// TIA Portal project "g" (V14) (continued)

   REGION Init
       IF #mb_query.z.run.state = #INIT_QUERY THEN
           // Modicon convention address conversion.
           "mb_internal_a"(mode104 := false,
                          Mode => #master.MODE,
                          Data_addr => #master.DATA_ADDR,
                          mb_query := #mb_query);
           // Copy buffer to a non optimiced memory area.
           IF #mb_query.z.run.write THEN
               #buffer.buffer := #mb_query.z.buffer;
           END_IF;
           // Automatically adjust timeout.
           #comm_load.RESP_TO := T_CONV
           (* *)("mb_timeout_rtu_calc"
                 (**)(gain := #conf.timeout_gain, 
                 (**) offset := #conf.timeout_offset,
                 (**) baud := #baud, mb_query := #mb_query));
           #comm_load.RETRIES := #conf.retries;
       END_IF;

       // Initiate the hardware
       #comm_load(REQ := #mb_query.z.run.state = #INIT_QUERY,
                  PORT := #hardware_id,
                  BAUD := #baud,
                  PARITY := #conf.parity, // Even is default.
                  RESP_TO := #comm_load.RESP_TO,
                  MB_DB := #master);

       IF #mb_query.z.run.state = #INIT_QUERY THEN
           IF #comm_load.DONE THEN
               #mb_query.z.run.state := #EXEC_QUERY;
           ELSE
               // Skip query exec. if init hw didn't go well.
               // The state RECIVE_RESUALT is inside mb_query.
               #mb_query.z.run.state := #RECIVE_RESUALT;
               #mb_query.stat.done := false;
               #mb_query.stat.error := true;
               #mb_query.stat.error_comm := true;
               #mb_query.stat.status := #comm_load.STATUS;
           END_IF;
       END_IF;
   END_REGION

   REGION Exec
       // The core master block.
       #master(REQ := #mb_query.z.run.state = #EXEC_QUERY
               AND NOT #master.BUSY,
               MB_ADDR := #mb_query.z.q.mb_addr,
               MODE := #master.MODE,
               DATA_ADDR := #master.DATA_ADDR,
               DATA_LEN := #mb_query.z.q.data_len,
               BUSY => #mb_query.stat.busy,
               DATA_PTR := #buffer.buffer);

       IF #mb_query.z.run.state = #EXEC_QUERY THEN
           #mb_query.stat.error := #master.ERROR;
           #mb_query.stat.done := #master.DONE;
           #mb_query.stat.status := #master.STATUS;
           "mb_internal_f"(buffer := #buffer, mb_query := #mb_query);
       END_IF;
   END_REGION

   // End is a comman FB for both tcp and rtu.
   #end(mb_query := #mb_query, Error => #Error);
END_FUNCTION_BLOCK

// folder: Library/Modbus/Core/Special

FUNCTION_BLOCK "mb_delay"   // FB11, SCL
{ S7_Optimized_Access := 'TRUE' }
VERSION : 0.1
   VAR_INPUT
      delay : Time;
   END_VAR
   VAR_IN_OUT
      mb_query : "mb_query";
   END_VAR
   VAR
      "timer" : TON_TIME;
      halt : Bool;
   END_VAR
BEGIN
   // For use with modbus tcp, so the client dosen't jam a network.
   // The function halt execution of queries for a certain time

   #mb_query.z.run.qid_cnt += 1;  // The timer occupy one qid.

   IF #halt // If the timer has been activated.
       OR #delay = T#0s // #delay = T#0s => Disable function
   THEN
       PRESET_TIMER(PT := #delay, TIMER := #"timer");
       #"timer"(IN := #delay <> T#0s, PT := #delay);
       IF #"timer".Q OR #delay = T#0s THEN
           IF #halt THEN
               #mb_query.conf.halt := #halt := false; // Continue exec.
               RESET_TIMER(#"timer");
           END_IF;
           #mb_query.z.run.qid += BOOL_TO_UINT
           (* *)(#mb_query.z.run.qid = #mb_query.z.run.qid_cnt);
       END_IF;

   ELSIF #mb_query.z.run.qid_cnt = #mb_query.z.run.qid THEN
       #mb_query.conf.halt := #halt := true; // Halt exec.
   END_IF;
END_FUNCTION_BLOCK

FUNCTION_BLOCK "mb_delay_between_queries"   // FB13, SCL
{ S7_Optimized_Access := 'TRUE' }
VERSION : 0.1
   VAR_INPUT
      delay : Time;
   END_VAR
   VAR_IN_OUT
      mb_query : "mb_query";
   END_VAR
   VAR
      "timer" : TON_TIME;
      halt : Bool;
      old_state : UInt;
   END_VAR
   VAR CONSTANT
      ORIGIN : USInt := 0;
   END_VAR
BEGIN
   // For use with modbus tcp, so the client dosen't jam a network.
   // The function halt execution of queries for a certain time
   // not just once, but between every query. There should only be
   // one of this block for each client.

   IF #halt // Is exec. halted?
       OR #delay = T#0s // #delay = T#0s => Disable function.
   THEN
       PRESET_TIMER(PT := #delay, TIMER := #"timer");
       #"timer"(IN := #delay <> T#0s, PT := #delay);
       IF #"timer".Q
           OR #delay = T#0s AND #halt
       THEN
           RESET_TIMER(#"timer");
           #mb_query.conf.halt := #halt := false; // Continue exec.
       END_IF;

   ELSIF #mb_query.z.run.state <> #old_state
       AND #mb_query.z.run.state <> #ORIGIN
   THEN
       // Halt exec. when next query is about to be inserted,
       // but current query will still finish.
       #mb_query.conf.halt := #halt := true; // Halt exec.
   END_IF;
   #old_state := #mb_query.z.run.state;
END_FUNCTION_BLOCK

FUNCTION "mb_query_bits" : Void   // FC9, SCL
{ S7_Optimized_Access := 'TRUE' }
VERSION : 0.1
   VAR_IN_OUT
      data_ptr : Array[*] of Bool;
      mb_query : "mb_query";
   END_VAR
   VAR_TEMP
      discrete : Bool;
      dommy : Bool;
      lower : DInt;
      upper : DInt;
      bits : UInt;
      bytes : UDInt;   // bytes
   END_VAR
   VAR CONSTANT
      INIT_QUERY : USInt := 2;
      RECIVE_RESUALT : USInt := 4;
   END_VAR
BEGIN
   // This function may be used when the number of bits dosen't
   // add up to whole bytes, for function codes: 1, 2, 5 and 15. 
   // 
   // data_ptr need to be a one dimensional array of bools.
   // --- --- ---

   REGION Header
       IF #mb_query.z.run.qid_cnt + 1 <> #mb_query.z.run.qid
           OR #mb_query.stat.busy
       THEN
           // Skip query, qid will not match qid_cnt and
           // my_query will return.
           #mb_query(data_ptr := #dommy);
           RETURN;
       END_IF;
   END_REGION

   REGION Pre-calc
       // Some preparing calculations.
       CASE #mb_query.mode OF // A discrete query ?
           1, 2, 5, 15:
               #discrete := true;
           200..202:
               CASE #mb_query.data_addr OF
                   1..19999: // 1..9999, 10001..19999
                       #discrete := true;
               END_CASE;
       END_CASE;
       #lower := LOWER_BOUND(ARR := #data_ptr, DIM := 1);
       #upper := UPPER_BOUND(ARR := #data_ptr, DIM := 1);
       #bits := DINT_TO_UINT(#upper - #lower + 1); // Elements in array.

       // Auto data len ?
       IF #mb_query.data_len = #mb_query.c.auto_len THEN
           #bytes := (#bits + 7) / 8; // CEIL()
           #mb_query.data_len := SEL(G := #discrete,
                                     IN0 := (#bits + 15) / 16, // CEIL()
                                     IN1 := #bits);
       ELSE
           #bytes := SEL(G := #discrete,
                         IN0 := #mb_query.data_len * 2, // 1 word -> 2 bytes
                         IN1 := (#mb_query.data_len + 7) / 8); // CEIL()
       END_IF;
   END_REGION

   REGION Run
       // Disable buf.h. inside mb_query.
       #mb_query.conf.buffer_handler := false;

       // Run the query.
       #mb_query(data_ptr := #dommy);

       #mb_query.conf.buffer_handler := true; // Enable buf.h. again.
       #mb_query.data_len := #mb_query.c.auto_len; // Back to auto.
   END_REGION

   REGION Insert & recive
       IF #mb_query.z.run.state = #INIT_QUERY  // Insert query.
           AND #mb_query.z.run.write
       THEN
           // Copy the content from data_ptr to the buffer.
           GATHER_BLK(IN := #data_ptr[#lower],
                      COUNT_OUT := #bytes,
                      OUT => #mb_query.z.buffer[0]);

       ELSIF  #mb_query.Done // The query above.
           AND NOT #mb_query.z.run.write  // A read query
       THEN
           // Copy the content from the buffer to data_ptr.
           SCATTER_BLK(IN := #mb_query.z.buffer[0],
                       COUNT_IN := #bytes,
                       OUT => #data_ptr[#lower]);
       END_IF;
   END_REGION
END_FUNCTION

// folder: Library/Modbus/Core/sb

FUNCTION "mb_station_block_header" : Void   // FC10, SCL
{ S7_Optimized_Access := 'TRUE' }
VERSION : 1.0
   VAR_IN_OUT
      sb : "mb_station_block_udt";
      mb_query : "mb_query";
   END_VAR
   VAR CONSTANT
      ORIGIN : USInt := 0;
   END_VAR
BEGIN
   // Rexhip - Extended modbus library.
   // Read the top section of mb_query for more documentation.

   // Skip everything !
   IF #sb.conf.skip_code THEN
       RETURN;
   END_IF;

   #mb_query.data_len := 0; // Default is auto-length.
   #mb_query.conf.buffer_handler := true;

   // If device blocks are executeded in diffrent order, a wide wind
   // up effect will occur, (in same OB) this will prevent that.
   IF #mb_query.z.sb.reset THEN
       #sb.z.header_qid := #mb_query.z.run.qid_cnt + 1;
   END_IF;

   // Device id cnt. The first device has id "1". Increased in every
   // mb_device_header, reseted in mb_client_ctrl or mb_master_ctrl.
   #mb_query.z.sb.sid_cnt += 1;

   // mb_query set the same bellow variables to true, at insert or recive.
   // This informastion is later used at the footer.
   #mb_query.z.sb.head_insert := false;
   #mb_query.z.sb.head_recive := false;

   // Reset order, a variable that makes queries in a sb execute in order.
   // #mb_query.z.sb.order := false;

   // When #mb.mb.q.qid = #mb.mb.run.qid_cnt => "This" device has the
   // query-token !
   // - If the query-token points at this device header, or it point to a
   //   query in the previous device, that is surrounded by a if-statement
   //   and the statement is now false.
   // - A gid change can only be done if not "busy", this is to avoid a
   //   resualt from one query being intercepted by another
   IF #mb_query.z.run.qid > #mb_query.z.run.qid_cnt
       AND #mb_query.z.run.qid <= #sb.z.header_qid
       AND NOT #mb_query.stat.busy
   THEN
       // Reset.
       // Go back to the first state in mb_query. New query param. will
       // owerwrite old once.
       #mb_query.z.run.state := #ORIGIN;

       // At first the offset_qid points at the first query of this
       // device. When it has executed the offset will point at the
       // second query. When all queries has executed the offset will
       // be reset back to the first query. (footer) 
       #mb_query.z.run.qid :=
       (* *)#sb.z.header_qid + #sb.z.offset_qid;

       // Order is a variable that makes queries in sb execute in order.
       //    #mb_query.z.sb.order := true;
   END_IF;

   // - The code below is reduce the impact of setting a if-statement
   //   around queries, by setting the qid_cnt to a fixed value at this 
   //   point.
   // - mb_station_block_header will occupy one query-id.  
   #sb.z.header_qid :=
   MAX(IN1 := #mb_query.z.run.qid_cnt + 1,
       IN2 := #sb.z.header_qid);
   #mb_query.z.run.qid_cnt := #sb.z.header_qid;
END_FUNCTION

FUNCTION "mb_station_block_footer" : Void   // FC11, SCL
{ S7_Optimized_Access := 'TRUE' }
VERSION : 1.0
   VAR_IN_OUT
      sb : "mb_station_block_udt";
      mb_query : "mb_query";
   END_VAR
   VAR_TEMP
      "e" : Int;
      err : Bool;
   END_VAR
   VAR CONSTANT
      INSERT_QUERY : USInt := 1;
   END_VAR
BEGIN
   // Rexhip - Extended modbus library.
   // Read the top section of mb_query for more documentation.

   // Skip everything !
   IF #sb.conf.skip_code THEN
       RETURN;
   END_IF;

   REGION Recive
       IF #mb_query.z.sb.head_recive THEN
           // If there is a query that bellong to this device that has
           // recvied a resault. (with or without error)

           // Counter for exec. queries inside this station block.
           // Default is 1 query for each loop, but may be changed.
           #sb.z.exec_cnt += 1;

           // If this is the first succesfylly query after communication error,
           // then log the time this happen. (also exceptions)
           IF #sb.out.error_comm AND (
               #mb_query.stat.done
               OR #mb_query.stat.error AND NOT #mb_query.stat.error_comm)
           THEN
               #"e" := RD_LOC_T(#sb.log.connected_time);
           END_IF;

           IF #mb_query.stat.error THEN // Logging - failed query        
               // Store the values for debugging. data_addr will indicate witch 
               // query caused the error, and the status is indicate the error type.
               #sb.log.error_status := #mb_query.stat.status;
               #sb.log.error_data_addr := #mb_query.z.sb.log_data_addr;

               // Two counters, one for comm.error and for all other errors.
               IF #mb_query.stat.error_comm THEN
                   #sb.log.error_comm_cnt += 1; // Eg. Bad CRC, parity, etc.
               ELSE
                   #sb.log.error_exception_cnt += 1;
               END_IF;

               // Increase communication error counter. if it's a comm.error.
               // then reset the counter.  
               IF #mb_query.stat.error_comm THEN
                   #sb.z.comm_err_cnt += BOOL_TO_USINT(#sb.z.comm_err_cnt < 255);
               ELSE
                   #sb.z.comm_err_cnt := 0;
               END_IF;

               // The error_comm flag is set if x repeating comm.errors occurres.
               #err := #sb.z.comm_err_cnt > #sb.conf.max_comm_error;
               IF #err AND NOT #sb.out.error_comm THEN
                   // Log the time when the flag is set.
                   #"e" := RD_LOC_T(#sb.log.disconnected_time);
               END_IF;
               #sb.out.error_comm := #err;

               // A comm.error will not be displayed before the
               // communication_error flag is set. Other errors will be
               // diplayed once. (NOT comm.error -> normal error)
               #sb.out.error := #sb.out.error OR NOT #mb_query.stat.error_comm
               OR #sb.out.error_comm;

               // err_hold makes the error flag stay true for more then just
               // one plc-scan.
               #sb.z.err_hold := #sb.out.error;

           ELSIF #mb_query.stat.done THEN // Logging successfully query        
               #sb.log.done_cnt += 1;
               // One successfully query -> reset fault.
               #sb.out.error_comm := false;
               #sb.z.comm_err_cnt := 0;
           END_IF;

           // - If it's this devices has the retry token, (sid_retry = sid_cnt)
           //   a retry has been executed and faild. Then set the retry_finished
           //   flag.
           // - The retry-token will be passed on to the next device with
           //   communication problems when the query loop has reach
           //   the end. (Inside the mb_internal_e)
           // - The library make sure that only one station block with comm.
           //   problems will do retry for each query loop revolution. 
           #mb_query.z.sb.retry_finished :=
           #mb_query.z.sb.sid_retry = #mb_query.z.sb.sid_cnt
           AND #mb_query.stat.error_comm;

           // Only one query in the SB is executed (default). The purpose is
           // to avoid a SB with many queries to occupy the bus for long periodes
           // of time. offset_qid is incread by one when a query has executed
           // given last query didn't resualt in a timeout.
           #sb.z.offset_qid += BOOL_TO_UINT(NOT #mb_query.stat.error_comm);
       END_IF;
   END_REGION

   REGION Middle
       // If all queries for this device has been executed,
       // then reset offset_qid back to the first query.
       IF #sb.z.offset_qid >
           #mb_query.z.run.qid_cnt - #sb.z.header_qid
       THEN
           #sb.z.offset_qid := 1;

           // Also reset error falg, if the last query was successfully.
           IF NOT #sb.z.err_hold THEN
               #sb.out.error := false;
           END_IF;
           #sb.z.err_hold := false;
       END_IF;

       // If the retry-token point at this device (sid_retry=sid_cnt), and there is
       // no communication problems then pass on the retry-token to the next device.
       // The retry token tell which device with communication problem that should
       // retry establish communication.
       #mb_query.z.sb.sid_retry +=
       BOOL_TO_UINT(#mb_query.z.sb.sid_retry = #mb_query.z.sb.sid_cnt
                    AND NOT #sb.out.error_comm);
   END_REGION

   REGION Finnish
       // Several condition that resault in passing on the query-token on to the
       // next device. Skipping all or the rest of the queries for this device:              
       #sb.out.finnish :=
       #mb_query.z.sb.head_recive AND ( // Skip rest of the queries if: ->
       (* *)#sb.z.exec_cnt >= #sb.conf.exec_x_quries // Some queries has executed,
       (*           *)// wait for the next loop for the remaining queries.
       (*      *)OR #mb_query.stat.error_comm) // A query resualting in comm.error    
       OR #mb_query.z.sb.head_insert AND ( // Erase a already inserted query if: ->
       (* *)#sb.out.error_comm // This station has allready comm. problems.
       (*      *)// And, it isn't this devies turn to try again.
       (*      *)AND (#mb_query.z.sb.sid_retry <> #mb_query.z.sb.sid_cnt
       (*           *)// Or, there has allready been a retry attempt on this loop.
       (*           *)OR #mb_query.z.sb.retry_finished) // (reseted in mb_internal_e)     
       (* *)OR #sb.conf.disable    
       (* *)OR #sb.conf.exec_x_quries = 0 // Zero => disable station block.
       (* *)OR #sb.conf.read_only // The read_only flag is set, and it's a write query.
       (*      *)AND #mb_query.z.run.write);

       IF #sb.out.finnish THEN // Reset
           // Go back to the first state in mb_query. New query param. will owerwrite 
           // old once.
           #mb_query.z.run.state := #INSERT_QUERY;
           // Set to qid to the next station block.
           #mb_query.z.run.qid := #mb_query.z.run.qid_cnt + 1;
           #sb.z.exec_cnt := 0;
       END_IF;
   END_REGION
END_FUNCTION

// folder: Library/Modbus/Core/z Internal

FUNCTION_BLOCK "mb_internal_b"   // FB6, SCL
{ S7_Optimized_Access := 'FALSE' }
VERSION : 0.1
   VAR
      buffer : Array[0..249] of Byte;
   END_VAR
BEGIN
   (*
   - Buffer for mb_master and modbus_master. (modbus rtu)
   - This block has optimize data access disabled.
   - For RTU, please do not delete the even there is no code bellow.
   - This block isn't needed for modbus tcp.
   *)
END_FUNCTION_BLOCK

FUNCTION_BLOCK "mb_internal_e"   // FB7, SCL
{ S7_Optimized_Access := 'TRUE' }
VERSION : 0.1
   VAR_OUTPUT
      Error : Bool;
   END_VAR
   VAR_IN_OUT
      mb_query : "mb_query";
   END_VAR
   VAR
      err_hold : Bool;
   END_VAR
   VAR CONSTANT
      INSERT_QUERY : USInt := 1;
      EXEC_QUERY : USInt := 3;
      RECIVE_RESUALT : USInt := 4;
   END_VAR
BEGIN
   // Internal function - common for both rtu and tcp.

   // Move on to next state when query is finnished.
   IF #mb_query.z.run.state = #EXEC_QUERY 
       AND (#mb_query.stat.error OR #mb_query.stat.done)
   THEN
       #mb_query.z.run.state := #RECIVE_RESUALT;
   END_IF;


   // Anti wind up effect for qid. msg. to devices that they should
   // reset if qid grow bigger then 60000. (See mb_station_block_header)
   #mb_query.z.sb.reset := false;
   IF #mb_query.z.run.qid > 60000 THEN
       #mb_query.z.sb.reset := true;
   END_IF;

   // #error will be keeped true as long there is at least one query that
   // generate a error. 
   IF #mb_query.stat.error THEN
       #Error := true;
       #err_hold := true;
   END_IF;

   // If all queries has been executed,
   IF #mb_query.z.run.qid > #mb_query.z.run.qid_cnt THEN

       // Error handeling (see above)
       IF NOT #err_hold THEN
           #Error := false;
       END_IF;
       #err_hold := false;

       // Start over again on the first query.
       #mb_query.z.run.qid := 1;

       // The retry-id is the device that get to have retry to restoring
       // communication after the error_comm flag is set for the station.
       // When one query loop has occurred the retry id is incremented. 
       #mb_query.z.sb.sid_retry := #mb_query.z.sb.sid_retry + 1;

       // retry_finished is set after one retry has taken place. 
       // The station that has the retry-token only has one try to make 
       // successfully query.
       #mb_query.z.sb.retry_finished := false;
       IF #mb_query.z.sb.sid_retry > #mb_query.z.sb.sid_cnt THEN
           #mb_query.z.sb.sid_retry := 1;
       END_IF;

       // Station id: (not in use)
       #mb_query.z.sb.sid := #mb_query.z.sb.sid + 1;
       IF #mb_query.z.sb.sid > #mb_query.z.sb.sid_cnt THEN
           #mb_query.z.sb.sid := 1;
       END_IF;
   END_IF;

   #mb_query.z.run.qid_cnt := 0; // (Incremented in mb_query)
   #mb_query.z.sb.sid_cnt := 0; // (Incremented in mb_station_block_header)
END_FUNCTION_BLOCK

FUNCTION "mb_internal_f" : Void   // FC2, SCL
{ S7_Optimized_Access := 'TRUE' }
VERSION : 0.1
   VAR_IN_OUT
      buffer : "mb_internal_b";
      mb_query : "mb_query";
   END_VAR
   VAR_TEMP
      comm_error : Bool;
   END_VAR
BEGIN
   // Internal function - master footer

   IF #mb_query.stat.error THEN
       // Figur out if it's a communication error.
       // (Handled different from other errors)
       CASE WORD_TO_UINT(#mb_query.stat.status) OF
           16#80C8, // Timeout
           16#80E1, // Parity error
           16#80E2, // Framing error
           16#8380: // Bad CRC 
               #comm_error := true;
       END_CASE;

   ELSIF #mb_query.stat.done // Successful query
       AND NOT #mb_query.z.run.write // A read query.
   THEN
       #mb_query.z.buffer := #buffer.buffer;
   END_IF;

   #mb_query.stat.error_comm :=
   (* *)#mb_query.stat.error AND #comm_error;
END_FUNCTION

FUNCTION "mb_internal_a" : Void   // FC4, SCL
{ S7_Optimized_Access := 'TRUE' }
VERSION : 0.1
   VAR_INPUT
      mode104 : Bool;
   END_VAR
   VAR_OUTPUT
      Mode : USInt;
      Data_addr : UDInt;
   END_VAR
   VAR_IN_OUT
      mb_query : "mb_query";
   END_VAR
BEGIN
   // Internal function

   // Modicon convention address.
   #Mode := 0;
   CASE #mb_query.z.q.mode OF
       1:  // Read output bits
           #Data_addr := 1 + #mb_query.z.q.data_addr;
       2:  // Read input bits
           #Data_addr := 10001 + #mb_query.z.q.data_addr;
       3:  // Read holding reg.
           #Data_addr := 400001 + #mb_query.z.q.data_addr;
       4:  // Read input word
           IF #mode104 THEN
               #Mode := 104;
               #Data_addr := #mb_query.z.q.data_addr;
           ELSE
               #Data_addr := 30001 + #mb_query.z.q.data_addr;
           END_IF;
       5:  // Writing a single output bit
           #Mode := 1;
           #Data_addr := 1 + #mb_query.z.q.data_addr;
       6:  // Writing a single holding register
           #Mode := 1;
           #Data_addr := 400001 + #mb_query.z.q.data_addr;
       15: // Writing multiple output bits
           #Mode := 2;
           #Data_addr := 1 + #mb_query.z.q.data_addr;
       16: // Writing multiple holding registers
           #Mode := 2;
           #Data_addr := 400001 + #mb_query.z.q.data_addr;
       200..202: // Read and write
           #Mode := #mb_query.z.q.mode - 200;
           #Data_addr := #mb_query.z.q.data_addr;
       ELSE
           #Mode := #mb_query.z.q.mode;
           #Data_addr := #mb_query.z.q.data_addr;
   END_CASE;
END_FUNCTION

FUNCTION "mb_timeout_rtu_calc" : Time   // FC5, SCL
{ S7_Optimized_Access := 'TRUE' }
VERSION : 0.1
   VAR_INPUT
      gain : Real;
      offset : Time;
      baud : UDInt;
   END_VAR
   VAR_IN_OUT
      mb_query : "mb_query";
   END_VAR
   VAR_TEMP
      t : Time;
   END_VAR
BEGIN
   // Automatically adjust timeout for modbus rtu.

   IF #gain = 0 THEN
       #t := #offset;
   ELSE
       #t := T_CONV
       (REAL_TO_UINT
        (
         11000 * ( //  11: Bits: start, data, parity, stop. 
         (* *)//   * 1000: Seconds to milliseconds
         (* *)19 // Bytes: Req: mb_addr, fc, data_addr(2), data_len(2), crc(2), 
         (* *) //        + res: mb_addr, fc, byte-count, crc(2), 
         (* *) //        + start-stop -> 6 (ca 2 x 28 bits)
         (* *)+ UINT_TO_REAL(#mb_query.z.q.data_len) *
         (*     *)SEL(G := #mb_query.z.run.discrete,
                      (* *)IN0 := INT_TO_REAL(2), // Each word is to bytes.
                      (* *)IN1 := 0.125) // Eight bits in one byte. (1/8 = 0.125)
         )
         / UDINT_TO_REAL(#baud) // High baud-rate -> low timeout
         * #gain // Safty margin
         + UDINT_TO_UINT(T_CONV(#offset))
        ));
   END_IF;

   #mb_timeout_rtu_calc :=
   LIMIT(MN := T#5ms, // A least 5ms, else comm_load will throw a error.
         IN := #t,
         MX := T#65s);
END_FUNCTION

// ===== library types =====

TYPE "timerUdt"
   STRUCT
      pt : Real;   // Preset time
      format : SInt := 2;   // 1=ms, 2=sec, 3=min, 4=h, 5=day
      RT : Real;   // Remaining time
   END_STRUCT;
END_TYPE

TYPE "ioGlobalUdt"
   STRUCT
      ackAllAlarms : Bool;   // Acknowledge all alarms
      disableAllSim : Bool;   // Disable all simulation of input values
      hmiShowTags : Bool;
      _ : Bool;
      totalActiveSim : UInt;   // Total active simulations
      totalActiveAlarms : UInt;   // Total active alarms
      totalUnacknowledgedAlarms : UInt;
      totalErrors : UInt;
   END_STRUCT;
END_TYPE

TYPE "alarmRealUdt"
   STRUCT
      value : Real;
      action : SInt;
      lim : Real;   // Alarm limit
      hyst : Real;   // Hysteresis
      delay : Time;   // Alarm delay
      delayEt : Time;   // delay elapsed time
      enable : Bool;   // Enable alarm
      autoAck : Bool := TRUE;   // manual acknowledge
      dobleAck : Bool;
      ack : Bool;   // acknowledge alarm
      memAck : Bool;   // Can be used for buzzer
      Q : Bool;   // output
   END_STRUCT;
END_TYPE

TYPE "analogInUdt"
   STRUCT
      filterConst : Real;   // 0=off , const for average filter.
      unitInterval : Real;   // 00.0 to 1.00 , (raw value, after running avg filter)
      sim : Bool;   // Simulate value
      forceInsideScale : Bool := true;   // Eg. in case of more then 20mA or less then 4mA.
      Error : Bool;   // Input signal out of range.
      zOldError : Bool;   // Internal variable
      ErrorTime : DTL;   // Time when the error occurred.
      errorAction : SInt := 100;   // [%]
      scaleMin : Real := 0.0;   // Scaled value for 4mA.
      scaleMax : Real := 100.0;   // Scaled value for 20mA.
      gain : Real := 1.0;   // Muliplied with the scaled value.
      offset : Real := 0.0;   // Added to "Q".
      Q : Real;   // value
   END_STRUCT;
END_TYPE

TYPE "analogInAndAlarmsUdt"
   STRUCT
      ai : "analogInUdt";
      execAiLogic : Bool := true;
      alarmL : "alarmRealUdt";
      alarmLL : "alarmRealUdt";
      alarmH : "alarmRealUdt";
      alarmHH : "alarmRealUdt";
      hmi : Struct
         copyAllSettings : Bool;
         pasteAllSettings : Bool;
         showTag : Bool;
      END_STRUCT;
   END_STRUCT;
END_TYPE

TYPE "alarmBoolSimpleUdt"
   STRUCT
      in : Bool;   // Input
      enable : Bool;   // Enable alarm
      autoAck : Bool := TRUE;   // Alarm will go away automaticaly when in goes false.
      dobleAck : Bool;
      ack : Bool;   // Acknowledge alarm
      memAck : Bool;   // Active alarm has been acknowledged
      Q : Bool;   // Output
   END_STRUCT;
END_TYPE

TYPE "digitalInUdt"
   STRUCT
      sim : Bool;   // Simulate input
      invert : Bool;   // Invert input
      Error : Bool;   // External error
      Q : Bool;   // Output
      delay : Time;   // Input delay
      delayEt : Time;
      alarm : "alarmBoolSimpleUdt";
      timeOn : DTL;
      timeOff : DTL;
   END_STRUCT;
END_TYPE

TYPE "intervalUdt"
   STRUCT
      time_between : Real;
      time_active : Real;
      time_format : SInt := 2;   // 1=ms, 2=sec, 3=min, 4=h, 5=day
      force_on : Bool;
      force_off : Bool;
      Q : Bool;
      RT : Real;
   END_STRUCT;
END_TYPE

TYPE "load_balancer_info_udt"
   STRUCT
      devices_in_operation : UInt;
      devices_standby : UInt;
      devices_started : UInt;
   END_STRUCT;
END_TYPE

TYPE "digitalOutUdt"
   STRUCT
      in : Bool;
      simEnable : Bool;
      simValue : Bool := 0;
      failSafe : Bool;
      failSafeValue : Bool;
      disableSim : Bool;
      invert : Bool;   // Invert output
   END_STRUCT;
END_TYPE

TYPE "timeFormatUdt"
   STRUCT
      OFF : SInt := 0;
      MILLISECOND : SInt := 1;
      SECOUNDS : SInt := 2;
      MINUTES : SInt := 3;
      HOURS : SInt := 4;
      DAYS : SInt := 5;
   END_STRUCT;
END_TYPE

TYPE "motorValveConfUdt"
   STRUCT
      toggleTimeBreak : Time := T#2S;   // A short break if valve change direction.
      regModeTimeBreak : Time := T#30S;   // Wait time before a new movment when valve is regMode
      regModeMinOffset : Real := 3.0;   // Min. offset before a movment is done when valve is in regMode.
      feilSafeAction : SInt := 2;   // 0=noAction, 1=open, 2=close.
      autoReset : Bool := TRUE;   // Reset on SP change or by jog valve, else iReset need to be set true.
      simFullyOpenWithPos : Bool;   // Use the pos-signal to determined if the valve is fully open.
      simFullyClosedWithPos : Bool;   // Use the pos-signal to determined if the valve is fully closed.
      fullyOpenPosLim : Real := 98.0;   // Above this position is seen as fully open
      fullyClosedPosLim : Real := 0.7;   // Under this position is seen as fully close
      gentleOpenEnable : Bool;   // Open valve with time breaks, this may prevent damange on equipment.
      gentleCloseEnable : Bool;   // Close valve with time breaks, this may prevent damange on equipment.
      gentleAlsoOnFailSafe : Bool := TRUE;   // The gentle function will also be enabled on fail safe mode.
      gentleActivteLowLimit : Real := 15.0;   // Gentle is only activate under this limit.
      gentleTimeRun : Time := T#2S_500MS;   // Valve movment time, on gentle open or close.
      gentleTimePauseBias : Real := 4.0;   // [s] Time break between each movment on gnetle open or close.
      gentleTimePauseDelta : Real := 20.0;   // [s] The time break will increase as fracton between limit and totaly closed.
      preStop : Real := 0.3;   // Stop the movment a bit before SP is reached, so the valve will stop exactly at SP.
      endPosWithoutPreStop : Real := 3.0;   // The few last procentages on close and open, there is no preStop
      longTimeout : Time := T#4M;   // If the valve hasn't reached it's position within this time, then there is something wrong.
      quickTimeoutEnable : Bool := TRUE;   // Check at interval that the valve move towards SP.
      quickTimeoutIntervalCheaks : Time := T#8S;   // Time interval between each check.
      qucikTimeoutMinMovement : Real := 2.0;   // Min movment between each check, else error.
   END_STRUCT;
END_TYPE

TYPE "operatingTimeUdt"
   STRUCT
      operatingTime : UDInt;
      startCnt : UDInt;
      oldIn : Bool;
      oldSec : USInt;
   END_STRUCT;
END_TYPE

TYPE "normXAnalogUdt"
   STRUCT
      rawMin : Int := 0;
      rawMax : Int := 27648;
      errorLimMin : Int := -4864;
      errorLimMax : Int := 32512;
   END_STRUCT;
END_TYPE

TYPE "pidUdt"
   STRUCT
      pidParam : PID_CompactControlParams;
      sp : Real;
      pv : Real;
      mv : Real;
      man : Bool;   // 0=auto
      error : Bool;
   END_STRUCT;
END_TYPE

// folder: Library/Alternating/Load balancer

TYPE "load_balancer_device_udt"
   STRUCT
      in_operation : Bool;   // Device in operation
      available : Bool := TRUE;   // Device is available for load balancer.
      Q : Bool;   // Main output
      operation_time : UDInt;   // sec
      z : Struct   // Internal variables
         n_cnt : UDInt;   // Used for boost start. (has nothing to do with this particular device)
      END_STRUCT;
   END_STRUCT;
END_TYPE

// folder: Library/Alternating/Load balancer/Blocks and UDT's

TYPE "load_balancer_settings_udt"
   STRUCT
      bypass : Bool;   // Setting bypass true make all outputs enabled.
      max_devices_same_time : UInt := 65535;   // Setting, max devices that can participate at the same time
      max_diff_operating : Struct   // Max operating time between device with most and least operating time
         sec : UDInt := 4_294_967_295;
         enable : Bool;
      END_STRUCT;
      start : Struct   // Condition for starting a device
         limit : Real := 90.0;
         delay : Time := T#3M;
         force : Bool;
      END_STRUCT;
      stop : Struct   // Condition for stopping a device
         limit : Real := 20.0;
         delay : Time := T#2M;
         force : Bool;
      END_STRUCT;
      info : Struct
         input : Real;   // Block input
         total : UInt;   // Total devices
         in_operation : UInt;   // Number of devices in operation
         standby : UInt;   // Devices standby for operation
         started : UInt;   // Devices started by load balancer.
      END_STRUCT;
      boostStart : Struct   // Start correct amout of devices right away.
         enable : Bool := true;
         auto : Bool := true;   // Based on statistic on how many is usually used.
         reset : Bool;   // Reset statistics about how many devices are most frequently running.
         devices : USInt;   // Number of devices to boost start
      END_STRUCT;
   END_STRUCT;
END_TYPE

// folder: Library/IO-handeling/Analog out

TYPE "analogOutUdt"
   STRUCT
      in : Real;   // Program input
      failSafe : Bool;
      interlook : Bool;
      simEnable : Bool;
      failSafeValue : SInt := 0;   // Percent value on error, -1=keep value
      scaleMin : Real := 0.0;
      scaleMax : Real := 100.0;   // (scaleMin=0)
      simValue : Real := 0.0;
   END_STRUCT;
END_TYPE

// folder: Library/Motor valve/Blocks and UDT's

TYPE "motorValveIoUdt"
   STRUCT
      in : Struct
         fullyOpen : Bool;
         fullyClosed : Bool;
         pos : Real;
         posError : Bool;
      END_STRUCT;
      out : Struct
         open : Bool;
         close : Bool;
      END_STRUCT;
      simulated : Bool;
   END_STRUCT;
END_TYPE

TYPE "motorValveHmiUdt"
   STRUCT
      conf : "motorValveConfUdt";
      io : "motorValveIoUdt";
      error : Struct
         timeout : Bool;
         posError : Bool;
      END_STRUCT;
      cmd : Struct
         reset : Bool;
         man : Bool;   // false=>auto
         auto : Bool;
         jogOpen : Bool;
         jogClose : Bool;
         openFully : Bool;
         closeFully : Bool;
         stop : Bool;
      END_STRUCT;
      info : Struct
         regMode : Bool;   // Most be activated if valve is controlled by a PID. Makes timebreaks between each move.
         failSafe : Bool;
         interlook : Bool;
      END_STRUCT;
      SP : Real;
      operatingTime : "operatingTimeUdt";
      sim : Struct   // Simulate feedback signal
         enable : Bool;
         pos : Real;
         simByPlc : Bool;
      END_STRUCT;
      autoMan : SInt := 2;
   END_STRUCT;
END_TYPE

// folder: (top level)

FUNCTION_BLOCK "digitalRippleFilter"   // FB1, SCL
{ S7_Optimized_Access := 'TRUE' }
VERSION : 0.1
   VAR_INPUT
      in : Bool;
      pt_on : Time;
      pt_off : Time;
   END_VAR
   VAR_OUTPUT
      Q : Bool;
   END_VAR
   VAR
      ton : TON_TIME;
      tof : TOF_TIME;
   END_VAR
BEGIN
   // Filter noice of a digital input signal.

   #ton(IN := #in, PT := #pt_on);

   #tof(IN := #ton.Q OR #tof.Q AND #in,
        PT := #pt_off,
        Q => #Q);
END_FUNCTION_BLOCK

FUNCTION_BLOCK "timerHmi"   // FB1, SCL
{ S7_Optimized_Access := 'TRUE' }
VERSION : 0.1
   VAR_INPUT
      in : Bool;   // Activate timer
      pt : Time;   // Added to internal "pt"
      TP : Bool;   // Puls timer
      TON : Bool;   // Timer-ON delay
      TOF : Bool;   // Timer-OFF delay
      TONR : Bool;   // Timer-ON retentiv.
   END_VAR
   VAR_OUTPUT
      Q : Bool;
      Error : Bool;   // More then one mode is active.
      RT : Time;
   END_VAR
   VAR_IN_OUT
      udt : "timerUdt";
   END_VAR
   VAR
      "timer" : IEC_TIMER;
   END_VAR
   VAR_TEMP
      p : Time;
   END_VAR
   VAR CONSTANT
      SECOUNDS : SInt;
   END_VAR
BEGIN
   // PT-max: 24 days, 20 hours, 31 min, 23 sec and 647 ms.
   // Format: 1=ms, 2=sec, 3=min, 4=h, 5=day

   // NOTE: #pt is add tho the interal preset time. (#tUdt.pt)
   #p := #pt + "real2time_format"(in := #udt.pt, format := #udt.format);

   #Error := 1 < // More then one mode is active?
   BOOL_TO_SINT(#TON) + BOOL_TO_SINT(#TOF) +
   BOOL_TO_SINT(#TP) + BOOL_TO_SINT(#TONR);

   IF #udt.format = 0 OR #Error THEN // Off
       RESET_TIMER(#"timer");
   ELSE
       // If pt is change while the timer has allread started then it will be
       // updated with the new preset time
       PRESET_TIMER(PT := #p, TIMER := #"timer");

       IF #TON THEN // Timer-ON delay
           #"timer".TON(IN := #in, PT := #p);
       ELSIF #TOF THEN // Timer-OFF delay
           #"timer".TOF(IN := #in, PT := #p);
       ELSIF #TP THEN // Puls timer
           #"timer".TP(IN := #in, PT := #p);
       ELSIF #TONR THEN // Timer-ON retentiv.
           #"timer".TONR(IN := #in, PT := #p);
       END_IF;
   END_IF;
   #Q := #"timer".Q;

   #RT := #p - #"timer".ET; // Remaining time.
   #udt.RT := "time2real_format"(in := #RT, format := #udt.format);
END_FUNCTION_BLOCK

FUNCTION_BLOCK "genUsrMsg"   // FB3, SCL
{ S7_Optimized_Access := 'TRUE' }
VERSION : 0.1
   VAR_INPUT
      TextID : UInt;
   END_VAR
   VAR
      TextListID : UInt;
      outgoingAlarm : Bool;   // false: Incoming alarm.
      assocValues : Array[3..10] of UInt;
      "e" : Int;
   END_VAR
   VAR_TEMP
      tmpAssocValues : AssocValues;
      c : Int;
   END_VAR
BEGIN
   // Generate user diagnostic alarms 

   // #assocValues 1 and 2 allready in use by instruction.
   FOR #c := 3 TO 10 DO
       #tmpAssocValues.Value[#c] := #assocValues[#c];
   END_FOR;

   #"e" := Gen_UsrMsg
   (Mode := 1 + BOOL_TO_UINT(#outgoingAlarm)
    ,// 1: incoming alarm. 2: outgoing alarm.
    TextID := #TextID,
   TextListID := #TextListID, // (Right click and show collom-id) 
    AssocValues := #tmpAssocValues);

   (* Assoc Values:

   "This is a usr. msg: @3I%6d@"  // Assoc val 3, 6 digits. (1st val)
   "This is an other usr. msg: @5I%6d@"  // Assoc val 5, 6 digits.

   *)
END_FUNCTION_BLOCK

FUNCTION_BLOCK "Interval"   // FB4, SCL
{ S7_Optimized_Access := 'TRUE' }
VERSION : 0.1
   VAR_INPUT
      in : Bool;   // Activate interval timer
   END_VAR
   VAR_OUTPUT
      Q : Bool;   // Output
      RT : Time;   // Remaining time
   END_VAR
   VAR_IN_OUT
      udt : "intervalUdt";
   END_VAR
   VAR
      N : UDInt;   // Number of cycles
      "timer" : IEC_TIMER;
   END_VAR
   VAR_TEMP
      r : Real;
      t : Time;
      "b" : Bool;
   END_VAR
   VAR CONSTANT
      SECOUNDS : SInt := 1;
   END_VAR
BEGIN
   // When #in is ture, then turn #Q on and off by preset times.

   #r := SEL(G := #udt.Q,
             IN0 := #udt.time_between,
             IN1 := #udt.time_active);
   #t := "real2time_format"(in := #r, format := #udt.time_format);
   PRESET_TIMER(PT := #t, TIMER := #"timer");
   #"timer".TON(IN := #in, PT := #t, Q => #"b");

   IF NOT #in THEN
       #udt.Q := false;
       #N := 0;
   ELSIF #udt.force_off THEN
       #udt.Q := false;
   ELSIF #udt.force_on THEN
       #udt.Q := true;
   ELSIF #"b" THEN
       #udt.Q := NOT #udt.Q; // Toggle.
       #N += BOOL_TO_UINT(#udt.Q);
   END_IF;

   IF #udt.force_off OR #udt.force_on OR #"b" THEN
       RESET_TIMER(#"timer");
       #udt.force_on := false;
       #udt.force_off := false;
   END_IF;

   #RT := #"timer".PT - #"timer".ET; // Remaining time
   #udt.RT := "time2real_format"(in := #RT, format := #udt.time_format);

   #Q := #udt.Q;
END_FUNCTION_BLOCK

FUNCTION_BLOCK "twoOutpus"   // FB5, SCL
{ S7_Optimized_Access := 'TRUE' }
VERSION : 0.1
   VAR_INPUT
      iStartOne : Bool;
      iStartBoth : Bool;
      iavailable1 : Bool := true;
      iavailable2 : Bool := true;
   END_VAR
   VAR_OUTPUT
      q1 : Bool;
      q2 : Bool;
   END_VAR
   VAR RETAIN
      next : SInt := 1;
   END_VAR
   VAR
      ftrig_in : F_TRIG;
   END_VAR
BEGIN
   // Alternating two outputs.

   #ftrig_in(CLK := #iStartOne);

   // Change #next if not available.
   IF NOT #iavailable1 AND #iavailable2 THEN
       #next := 2;
   ELSIF NOT #iavailable2 AND #iavailable1 THEN
       #next := 1;

   // Swap which one to start next time.
   ELSIF #ftrig_in.Q AND NOT #iStartBoth THEN
       #next := SEL(G := #next = 1,
                    IN0 := 1, IN1 := 2);

   // Make sure that value is valid, 1 or 2.    
   ELSIF #next <> 1 AND #next <> 2 THEN
       #next := 1;
   END_IF;

   #q1 := (#next = 1 AND #iStartOne OR #iStartBoth) AND #iavailable1;
   #q2 := (#next = 2 AND #iStartOne OR #iStartBoth) AND #iavailable2;
END_FUNCTION_BLOCK

FUNCTION_BLOCK "example_genUsrMsg"   // FB8, SCL
{ S7_Optimized_Access := 'TRUE' }
VERSION : 0.1
   VAR
      Gen_UsrMsg : "Gen_UsrMsg";
      some_error : Bool;
   END_VAR
BEGIN
   #Gen_UsrMsg.TextListID := 512; // See PLC alarm text lists.

   IF #some_error THEN
       #Gen_UsrMsg(1); // Text id for this alarm 
   END_IF;
END_FUNCTION_BLOCK

FUNCTION_BLOCK "motorValveAproxPos"   // FB8, SCL
{ S7_Optimized_Access := 'TRUE' }
VERSION : 0.1
   VAR_IN_OUT
      io : "motorValveIoUdt";
   END_VAR
   VAR
      conf : Struct
         maxAvoid : Real := 4.0;
      END_STRUCT;
      oldSecAndMsec10 : UInt;
      posPrT : UInt;
      "timer" : IEC_TIMER;
      first_scan : Bool := TRUE;
      RTRIG_fullyOpen : R_TRIG;
      RTRIG_fullyClosed : R_TRIG;
      rangeTime : Time;
      tries : Array[0..7] of Time;
   END_VAR
   VAR_TEMP
      "e" : Int;
      rd_sys_t : DTL;
      secAndMsec10 : UInt;
      sPos : Int;
      t : Int;
      c : Int;
      mx : Time;
      mn : Time;
   END_VAR
BEGIN
   // #io - "motorValveIoUdt"


   // For valve without position sensor. Calculate the position based on long
   // time the valve has been opening and closing.

   (* FUNCTION NOT FINISHED...

   #e := RD_SYS_T(#rd_sys_t);
   #secAndMsec10 := #rd_sys_t.SECOND * 100 + UDINT_TO_UINT(#rd_sys_t.NANOSECOND / 10000);
   #t := USINT_TO_INT( (#secAndMsec10 - #oldSecAndMsec10 + 6000) MOD 6000);
   #oldSecAndMsec10 := #secAndMsec10;

   #io.in.posError := #io.in.posError AND NOT #first_scan;

   #RTRIG_fullyOpen(CLK := #io.in.fullyOpen);
   #RTRIG_fullyClosed(CLK := #io.in.fullyClosed);

   IF #RTRIG_fullyOpen.Q OR #RTRIG_fullyClosed.Q THEN
       RESET_TIMER(#timer);
       #timer.PT := T#10m;
   END_IF;



   #c := 7 - 1;
   WHILE #c >= 0 DO
       #tries[#c + 1] := #tries[#c];
       #c -= 1;
   END_WHILE;
   #tries[0] := T#123s;

   #mn := T#24d;
   FOR #c := 1 TO 6 BY 2 DO
       #mx := MAX(IN1 := #tries[#c], IN2 := #mx);
       #mn := MIN(IN1 := #tries[#c], IN2 := #mn);
   END_FOR;
   // #mx - #mn ;

   (*IF #first_scan THEN
       #io.in.posError := true;
   END_IF;*)


   IF #io.out.open XOR #io.out.close THEN
       #sPos := SEL(G := #io.out.close, IN0 := #sPos + #t, IN1 := #sPos - #t);
   END_IF;


   // #io.in.pos

   #first_scan := false;

   *)
END_FUNCTION_BLOCK

FUNCTION_BLOCK "motorValveDigital"   // FB11, SCL
{ S7_Optimized_Access := 'TRUE' }
VERSION : 0.1
   VAR_INPUT
      iAction : SInt;   // 0=no-action, 1=Open, 2=Close
      iFailSafe : Bool;   // Open or close the valve entirly, set inside conf.
      iInterlook : Bool;   // Stop movement, valve will continue when input is set back false.
      iStop : Bool;   // Stop movement, also after var. is back false.
      iJogOpen : Bool;   // Move the valve towards open when true, has priority over SP.
      iJogClose : Bool;   // Move the valve towards close when true, has priority over SP.
      iReset : Bool;   // Reset timeout.
   END_VAR
   VAR_OUTPUT
      qTimeout : Bool;   // (quick and long timeout)
   END_VAR
   VAR
      action : SInt;   // 1=open, 2=close
      actionOut : SInt;
      oldAction : SInt;
      oldActionOut : SInt;
      RTIRG_iFailSafe : R_TRIG;
      RTIRG_iReset : R_TRIG;
      RTIRG_jog : R_TRIG;
      TP_toggleOut : IEC_TIMER;
      TON_gentle : IEC_TIMER;
      TONR_gentle : IEC_TIMER;
      TONR_timeout : IEC_TIMER;
      TON_regModeWait : IEC_TIMER;
      gentleAction : Bool;
   END_VAR
   VAR_TEMP
      reset : Bool;
   END_VAR
   VAR CONSTANT
      NO_ACTION : SInt := 0;
      OPEN : SInt := 1;
      CLOSE : SInt := 2;
   END_VAR
BEGIN
   // #conf - "motorValveConfUdt"
   // #io - "motorValveIoUdt"

   // Valve 

   (*

   //R-TRIG'S
   #RTIRG_iReset(CLK := #iReset);
   #RTIRG_iFailSafe(CLK := #iFailSafe); // Reset timeout once on failSafe.
   #RTIRG_jog(CLK := #iJogOpen XOR #iJogClose);

   REGION Timeout-and-reset
       // Max time the valve can operate before timeout, and the valve will stop.
       #TONR_timeout.TONR(IN := #io.out.open OR #io.out.close,
                          PT := #conf.longTimeout,
                          Q => #qTimeout);

       // Reset timeout
       IF #iJogOpen OR #iJogClose THEN
           #reset := #RTIRG_jog.Q AND (#conf.autoReset OR NOT #qTimeout);
       END_IF;
       IF #RTIRG_iReset.Q OR #RTIRG_iFailSafe.Q OR #reset THEN
           RESET_TIMER(#TONR_timeout);
           #qTimeout := false;
       END_IF;
   END_REGION

   REGION Decide
       // Error, timeout, failSafe and Interlook.
       IF #TONR_timeout.Q THEN
           #action := #NO_ACTION;
       ELSIF #iFailSafe THEN // Timeout will be reseted once if iFailSafe is activated.
           #action := #conf.feilSafeAction;
       ELSIF #iStop THEN
           #action := #NO_ACTION;
           // ==========================================================================
           // JOG-mode
       ELSIF #iJogOpen OR #iJogClose THEN
           // Open or close the valve little by little. When either of the jog
           // inputs are true. This way of controlling the valve has priority
           // over setpoint (bellow).
           RESET_TIMER(#TON_regModeWait);
           IF #iJogOpen AND #iJogClose THEN
               #action := #NO_ACTION;
           ELSIF #iJogOpen THEN
               #action := #OPEN;
           ELSIF #iJogClose THEN
               #action := #CLOSE;
           ELSE
               ;
           END_IF;
       END_IF;
   END_REGION

   REGION Gentle
       // If a big valve closes or open to fast, it can damage the pipes or other
       // equipment. This section make time breaks on closing or opening. 
       IF #io.in.pos < #conf.gentleActivteLowLimit // ->
           // -> The function is only active under a ceratain position limit.
           AND (NOT #iFailSafe OR #conf.gentleAlsoOnFailSafe)
           // AlsoOnFailSafe: It's possible to disable the function for emergencies
           // by setting the value false.
           AND (#conf.gentleOpenEnable AND #action = #OPEN
           (* *)OR #conf.gentleOpenEnable AND #action = #CLOSE)
       THEN
           #TON_gentle.PT := SEL(G := #gentleAction, // Toggle times
                                 IN0 := #conf.gentleTimeRun,
                                 IN1 := #conf.gentleTimePauseBias);
           #TON_gentle.TON(IN := true,
                           PT := #TON_gentle.PT);
           IF #TON_gentle.Q THEN
               #gentleAction := NOT #gentleAction;
               RESET_TIMER(#TON_gentle);
           END_IF;
           #actionOut := SEL(G := #gentleAction, // Toggle action
                             IN0 := #action, IN1 := #NO_ACTION);
       ELSE
           RESET_TIMER(#TON_gentle);
           #gentleAction := false;
           // If the carefully-function is disabled, then just forward
           // the action value to the next stage.
           #actionOut := #action;
       END_IF;
   END_REGION

   REGION Output
       // Make a smal time break when valve change direction. This make sure that
       // that both outputs are not active at the same time.
       #TP_toggleOut.TP(IN := #actionOut <> #oldActionOut AND #oldActionOut <> #NO_ACTION,
                        PT := #conf.toggleTimeBreak);
       // Outputs
       IF #TP_toggleOut.Q THEN
           #io.out.open := false;
           #io.out.close := false;
       ELSIF #iFailSafe THEN
           #io.out.open := #conf.feilSafeAction = #OPEN AND NOT #io.in.fullyOpen;
           #io.out.close := #conf.feilSafeAction = #CLOSE AND NOT #io.in.fullyClosed;
       ELSIF #iInterlook OR #iStop THEN
           #io.out.open := false;
           #io.out.close := false;
       ELSE
           #io.out.open := #actionOut = #OPEN AND NOT #io.in.fullyOpen;
           #io.out.close := #actionOut = #CLOSE AND NOT #io.in.fullyClosed;
       END_IF;
   END_REGION

   REGION Old
       #oldAction := #action;
       #oldActionOut := #actionOut;
   END_REGION


   // *)
END_FUNCTION_BLOCK

FUNCTION_BLOCK "_example_motorValve"   // FB12, SCL
{ S7_Optimized_Access := 'TRUE' }
VERSION : 0.1
   VAR_INPUT
      ai_valve1Pos : Int;
      di_valve1FullyOpen : Bool;
      di_valve1FullyClosed : Bool;
   END_VAR
   VAR_OUTPUT
      do_valve1Open : Bool;
      do_valve1Close : Bool;
   END_VAR
   VAR_IN_OUT
      ioGlobal : "ioGlobal_FB";
   END_VAR
   VAR
      valve1 : "motorValve";
      valve2 : "motorValve";
      motorValveSimulation_1 : "motorValveSimulation";
      motorValveSimulation_2 : "motorValveSimulation";
      speed : Real := 1.0;
   END_VAR
BEGIN

   // Valve 1 - (The linking block isn't required)
   "ioGlobalMotorValveLinking"(ioGlobal := #ioGlobal, valve := #valve1);
   #valve1
   (
    iFeedbackPosition := "analogInSimple"(mn := 0, in := #ai_valve1Pos, mx := 100),
    iFeddbackPosError := "analogInError"(#ai_valve1Pos),
    iFeedbackFullyOpen := #di_valve1FullyOpen,
    iFeedbackFullyClosed := #di_valve1FullyClosed,
    qOpen => #do_valve1Open,
    qClose => #do_valve1Close
   );

   // Vavle 2
   "ioGlobalMotorValveLinking"(ioGlobal := #ioGlobal, valve := #valve2);
   #valve2();

